FUNCTION_BLOCK "Connect"   // FB11, SCL
{ S7_Optimized_Access := 'TRUE' }
VERSION : 0.1
   VAR_INPUT
      tcon_param : TCON_Param;
   END_VAR
   VAR_IN_OUT
      requests : "Connection_Requests.UDT";
      saved_status : "Connection_Status.UDT";
   END_VAR
   VAR
      busy_delay_timer : TOF_TIME;
      error_timer : TOF_TIME;
      status_timer : TOF_TIME;
      TCON : TCON;
   END_VAR
   VAR_TEMP
      _block_status : "Connection_Status.UDT";
   END_VAR
BEGIN
   #TCON(REQ := #requests.connect,
         ID := #tcon_param.ID,
         DONE => #_block_status.done,
         BUSY => #_block_status.busy,
         ERROR => #_block_status.error,
         STATUS => #_block_status.status,
         CONNECT := #tcon_param);
   #requests.connect := FALSE;
   "Connect_Status.to_Control_Element"(requests := #requests,
                                          block_status := #_block_status,
                                          busy_timer := #busy_delay_timer,
                                          error_timer := #error_timer,
                                          saved_status := #saved_status,
                                          status_timer := #status_timer);
END_FUNCTION_BLOCK

// folder: tcpip_connection/connect/connect_status

FUNCTION "Connect_Status.Done" : Void   // FC138, SCL
{ S7_Optimized_Access := 'TRUE' }
VERSION : 0.1
   VAR_INPUT
      requests : "Connection_Requests.UDT";
      block_status : "Connection_Status.UDT";
   END_VAR
   VAR_IN_OUT
      saved_status : "Connection_Status.UDT";
   END_VAR
BEGIN
   "Connect_Status.Set_Done"(block_status := #block_status,
                                requests := #requests,
                                saved_status := #saved_status);
   "Connect_Status.Reset_Done"(block_status := #block_status,
                                  requests := #requests,
                                  saved_status := #saved_status);
END_FUNCTION

FUNCTION "Connect_Status.Error" : Void   // FC139, SCL
{ S7_Optimized_Access := 'TRUE' }
VERSION : 0.1
   VAR_INPUT
      block_status : "Connection_Status.UDT";
      requests : "Connection_Requests.UDT";
   END_VAR
   VAR_IN_OUT
      off_delay : TOF_TIME;
      saved_status : "Connection_Status.UDT";
   END_VAR
BEGIN
   "Connect_Status.Set_Error"(block_status := #block_status,
                                 requests := #requests,
                                 off_delay := #off_delay,
                                 saved_status := #saved_status);
END_FUNCTION

FUNCTION "Connect_Status.Reset_Busy" : Void   // FC140, SCL
{ S7_Optimized_Access := 'TRUE' }
VERSION : 0.1
   VAR_INPUT
      requests : "Connection_Requests.UDT";
   END_VAR
   VAR_IN_OUT
      saved_status : "Connection_Status.UDT";
   END_VAR
BEGIN
   IF #requests.disconnect THEN
       #saved_status.busy := FALSE;
   END_IF;
END_FUNCTION

FUNCTION "Connect_Status.Set_Busy" : Void   // FC142, SCL
{ S7_Optimized_Access := 'TRUE' }
VERSION : 0.1
   VAR_INPUT
      block_status : "Connection_Status.UDT";
      requests : "Connection_Requests.UDT";
   END_VAR
   VAR_IN_OUT
      off_delay : TOF_TIME;
      saved_status : "Connection_Status.UDT";
   END_VAR
   VAR_TEMP
      _et : Time;
   END_VAR
   VAR CONSTANT
      DELAY : Time := t#3s;
   END_VAR
BEGIN
   #off_delay(IN := #block_status.busy AND NOT #requests.disconnect,
              PT := #DELAY,
              Q => #saved_status.busy,
              ET => #_et);
END_FUNCTION

FUNCTION "Connect_Status.Busy" : Void   // FC143, SCL
{ S7_Optimized_Access := 'TRUE' }
VERSION : 0.1
   VAR_INPUT
      block_status : "Connection_Status.UDT";
      requests : "Connection_Requests.UDT";
   END_VAR
   VAR_IN_OUT
      off_delay : TOF_TIME;
      saved_status : "Connection_Status.UDT";
   END_VAR
BEGIN
   "Connect_Status.Set_Busy"(block_status := #block_status,
                                requests := #requests,
                                off_delay := #off_delay,
                                saved_status := #saved_status);
   "Connect_Status.Reset_Busy"(requests := #requests,
                                  saved_status := #saved_status);
END_FUNCTION

FUNCTION "Connect_Status.to_Control_Element" : Void   // FC144, SCL
{ S7_Optimized_Access := 'TRUE' }
VERSION : 0.1
   VAR_INPUT
      requests : "Connection_Requests.UDT";
      block_status : "Connection_Status.UDT";
   END_VAR
   VAR_IN_OUT
      busy_timer : TOF_TIME;
      error_timer : TOF_TIME;
      saved_status : "Connection_Status.UDT";
      status_timer : TOF_TIME;
   END_VAR
BEGIN
   "Connect_Status.Busy"(block_status := #block_status,
                            requests := #requests,
                            off_delay := #busy_timer,
                            saved_status := #saved_status);
   "Connect_Status.Done"(requests := #requests,
                            block_status := #block_status,
                            saved_status := #saved_status);
   "Connect_Status.Error"(block_status := #block_status,
                             requests := #requests,
                             off_delay := #error_timer,
                             saved_status := #saved_status);
   "Connect_Status.Status"(block_status := #block_status,
                              requests := #requests,
                              saved_status := #saved_status,
                              status_timer := #status_timer);
END_FUNCTION

FUNCTION "Connect_Status.Set_Done" : Void   // FC145, SCL
{ S7_Optimized_Access := 'TRUE' }
VERSION : 0.1
   VAR_INPUT
      block_status : "Connection_Status.UDT";
      requests : "Connection_Requests.UDT";
   END_VAR
   VAR_IN_OUT
      saved_status : "Connection_Status.UDT";
   END_VAR
BEGIN
   IF #block_status.done THEN
       #saved_status.done := TRUE;
   END_IF;
END_FUNCTION

FUNCTION "Connect_Status.Reset_Done" : Void   // FC146, SCL
{ S7_Optimized_Access := 'TRUE' }
VERSION : 0.1
   VAR_INPUT
      block_status : "Connection_Status.UDT";
      requests : "Connection_Requests.UDT";
   END_VAR
   VAR_IN_OUT
      saved_status : "Connection_Status.UDT";
   END_VAR
BEGIN
   IF #requests.disconnect THEN
       #saved_status.done := FALSE;
   END_IF;
END_FUNCTION

FUNCTION "Connect_Status.Set_Error" : Void   // FC147, SCL
{ S7_Optimized_Access := 'TRUE' }
VERSION : 0.1
   VAR_INPUT
      block_status : "Connection_Status.UDT";
      requests : "Connection_Requests.UDT";
   END_VAR
   VAR_IN_OUT
      off_delay : TOF_TIME;
      saved_status : "Connection_Status.UDT";
   END_VAR
   VAR_TEMP
      _et : Time;
   END_VAR
   VAR CONSTANT
      DELAY : Time := t#30s;
   END_VAR
BEGIN
   #off_delay(IN := #block_status.error,
              PT := #DELAY,
              Q => #saved_status.error,
              ET => #_et);
END_FUNCTION

FUNCTION "Connect_Status.Save_Status" : Void   // FC148, SCL
{ S7_Optimized_Access := 'TRUE' }
VERSION : 0.1
   VAR_INPUT
      block_status : "Connection_Status.UDT";
   END_VAR
   VAR_IN_OUT
      saved_status : "Connection_Status.UDT";
      status_timer : TOF_TIME;
   END_VAR
   VAR_TEMP
      _delay_update : Bool;
      _et : Time;
   END_VAR
   VAR CONSTANT
      DELAY : Time := T#30S;
      IDLE : Word := 16#7000;
   END_VAR
BEGIN
   IF #block_status.status <> #IDLE THEN
       #saved_status.status := #block_status.status;
   END_IF;
   #status_timer(IN := #block_status.status <> #IDLE,
                 PT := #DELAY,
                 Q => #_delay_update,
                 ET => #_et);
   IF #_delay_update THEN
       RETURN;
   END_IF;
   #saved_status.status := #block_status.status;
END_FUNCTION

FUNCTION "Connect_Status.Status" : Void   // FC149, SCL
{ S7_Optimized_Access := 'TRUE' }
VERSION : 0.1
   VAR_INPUT
      block_status : "Connection_Status.UDT";
      requests : "Connection_Requests.UDT";
   END_VAR
   VAR_IN_OUT
      saved_status : "Connection_Status.UDT";
      status_timer : TOF_TIME;
   END_VAR
BEGIN
   "Connect_Status.Save_Status"(block_status := #block_status,
                                   saved_status := #saved_status,
                                   status_timer := #status_timer);
   "Connect_Status.Clear_Status"(requests := #requests,
                                    saved_status := #saved_status);
END_FUNCTION

FUNCTION "Connect_Status.Clear_Status" : Void   // FC150, SCL
{ S7_Optimized_Access := 'TRUE' }
VERSION : 0.1
   VAR_INPUT
      requests : "Connection_Requests.UDT";
   END_VAR
   VAR_IN_OUT
      saved_status : "Connection_Status.UDT";
   END_VAR
BEGIN
   IF #requests.disconnect THEN
       #saved_status.status := 0;
   END_IF;
END_FUNCTION

// folder: tcpip_connection/connection_control

FUNCTION "Connection_Control.Initialize_Display" : Void   // FC85, SCL
{ S7_Optimized_Access := 'TRUE' }
VERSION : 0.1
   VAR_IN_OUT
      interface : "Connection_Status.HMI.UDT";
   END_VAR
BEGIN
   "Screen_Background.Initialize_Color"(#interface.background);
   "Screen_Background.Initialize_Visibility"(#interface.background);
   "Connection_Control_Table.Initialize_Display"(#interface.wire);
   "Connection_Control_Table.Initialize_Display"(#interface.material);
END_FUNCTION

// folder: tcpip_connection/connection_control/connection_control_element

FUNCTION "Connection_Control_Element.Initialize_Display" : Void   // FC86, SCL
{ S7_Optimized_Access := 'TRUE' }
VERSION : 0.1
   VAR_IN_OUT
      connection_status_element : "Connection_Status_Element.UDT";
   END_VAR
BEGIN
   "Connection_Control_Element.Initialize_Colors"(#connection_status_element);
   "Connection_Control_Element.Initialize_Visible"(#connection_status_element);
   "Connection_Control_Element.Initialize_Enable"(#connection_status_element);
END_FUNCTION

FUNCTION "Connection_Control_Element.Initialize_Colors" : Void   // FC87, SCL
{ S7_Optimized_Access := 'TRUE' }
VERSION : 0.1
   VAR_IN_OUT
      connection_status_element : "Connection_Status_Element.UDT";
   END_VAR
BEGIN
   #connection_status_element.busy_status_indicator_animate := "Color.String_to_DInt"("BUSY_INDICATOR_OFF");
   #connection_status_element.done_status_indicator_animate := "Color.String_to_DInt"("DONE_INDICATOR_OFF");
   #connection_status_element.error_status_indicator_animate := "Color.String_to_DInt"("ERROR_INDICATOR_OFF");
   #connection_status_element.operation_label_animate := "Color.String_to_DInt"("OPERATION_LABEL_OFF");
   #connection_status_element.status_code_description_animate := "Color.String_to_DInt"("STATUS_CODE_OFF");
   #connection_status_element.status_code_label_animate := "Color.String_to_DInt"("STATUS_CODE_OFF");
   #connection_status_element.status_code_value_animate := "Color.String_to_DInt"("STATUS_CODE_OFF");
END_FUNCTION

FUNCTION "Connection_Control_Element.Initialize_Visible" : Void   // FC88, SCL
{ S7_Optimized_Access := 'TRUE' }
VERSION : 0.1
   VAR_IN_OUT
      connection_status_element : "Connection_Status_Element.UDT";
   END_VAR
BEGIN
   #connection_status_element.busy_status_indicator_visible := TRUE;
   #connection_status_element.done_status_indicator_visible := TRUE;
   #connection_status_element.error_status_indicator_visible := TRUE;
   #connection_status_element.operation_button_visible := TRUE;
   #connection_status_element.operation_label_visible := TRUE;
   #connection_status_element.show_status_code_description_button_visible := TRUE;
   #connection_status_element.status_code_description_visible := TRUE;
   #connection_status_element.status_code_label_visible := TRUE;
   #connection_status_element.status_code_value_visible := TRUE;
END_FUNCTION

FUNCTION "Connection_Control_Element.Initialize_Enable" : Void   // FC89, SCL
{ S7_Optimized_Access := 'TRUE' }
VERSION : 0.1
   VAR_IN_OUT
      connection_status_element : "Connection_Status_Element.UDT";
   END_VAR
BEGIN
   #connection_status_element.operation_button_enable := TRUE;
   #connection_status_element.show_status_code_description_button_enable := TRUE;
END_FUNCTION

FUNCTION "Connection_Control_Element.Animate_Done" : Void   // FC94, SCL
{ S7_Optimized_Access := 'TRUE' }
VERSION : 0.1
   VAR_INPUT
      status : "Connection_Status.UDT";
   END_VAR
   VAR_IN_OUT
      interface : "Connection_Status_Element.UDT";
   END_VAR
BEGIN
   "Bool.Animate"(signal := #status.done,
                  color_on := "Color.String_to_DInt"("DONE_INDICATOR_ON"),
                  color_off := "Color.String_to_DInt"("DONE_INDICATOR_OFF"),
                  animation := #interface.done_status_indicator_animate);
END_FUNCTION

FUNCTION "Connection_Control_Element.Animate_Error" : Void   // FC95, SCL
{ S7_Optimized_Access := 'TRUE' }
VERSION : 0.1
   VAR_INPUT
      status : "Connection_Status.UDT";
   END_VAR
   VAR_IN_OUT
      interface : "Connection_Status_Element.UDT";
   END_VAR
BEGIN
   "Bool.Animate"(signal := #status.error,
                  color_on := "Color.String_to_DInt"("ERROR_INDICATOR_ON"),
                  color_off := "Color.String_to_DInt"("ERROR_INDICATOR_OFF"),
                  animation := #interface.error_status_indicator_animate);
END_FUNCTION

FUNCTION "Connection_Control_Element.Animate_Status_Bad" : Void   // FC96, SCL
{ S7_Optimized_Access := 'TRUE' }
VERSION : 0.1
   VAR_IN_OUT
      connection_status_element : "Connection_Status_Element.UDT";
   END_VAR
BEGIN
   #connection_status_element.status_code_description_animate := "Color.String_to_DInt"("STATUS_CODE_PROBLEM");
   #connection_status_element.status_code_label_animate := "Color.String_to_DInt"("STATUS_CODE_PROBLEM");
   #connection_status_element.status_code_value_animate := "Color.String_to_DInt"("STATUS_CODE_PROBLEM");
END_FUNCTION

FUNCTION "Connection_Control_Element.Animate_Busy" : Void   // FC97, SCL
{ S7_Optimized_Access := 'TRUE' }
VERSION : 0.1
   VAR_INPUT
      status : "Connection_Status.UDT";
   END_VAR
   VAR_IN_OUT
      element : "Connection_Status_Element.UDT";
   END_VAR
BEGIN
   "Bool.Animate"(signal := #status.busy,
                  color_on := "Color.String_to_DInt"("BUSY_INDICATOR_ON"),
                  color_off := "Color.String_to_DInt"("BUSY_INDICATOR_OFF"),
                  animation := #element.busy_status_indicator_animate);
END_FUNCTION

FUNCTION "Connection_Control_Element.Animate_Status_Good" : Void   // FC98, SCL
{ S7_Optimized_Access := 'TRUE' }
VERSION : 0.1
   VAR_IN_OUT
      interface : "Connection_Status_Element.UDT";
   END_VAR
BEGIN
   #interface.status_code_description_animate := "Color.String_to_DInt"("STATUS_CODE_GOOD");
   #interface.status_code_label_animate := "Color.String_to_DInt"("STATUS_CODE_GOOD");
   #interface.status_code_value_animate := "Color.String_to_DInt"("STATUS_CODE_GOOD");
END_FUNCTION

FUNCTION "Connection_Control_Element.Animate_Operation_Acutate" : Void   // FC135, SCL
{ S7_Optimized_Access := 'TRUE' }
VERSION : 0.1
   VAR_IN_OUT
      interface : "Connection_Status_Element.UDT";
   END_VAR
   VAR_TEMP
      _animation : DInt;
   END_VAR
BEGIN
   "Bool.Animate"(signal := #interface.operation_button_actuate,
                  color_on := "Color.String_to_DInt"("ACTUATE"),
                  color_off := "Color.String_to_DInt"("OPERATION_OFF"),
                  animation := #interface.operation_label_animate);
END_FUNCTION

FUNCTION "Connection_Control_Element.Animate" : Void   // FC141, SCL
{ S7_Optimized_Access := 'TRUE' }
VERSION : 0.1
   VAR_INPUT
      status : "Connection_Status.UDT";
   END_VAR
   VAR_IN_OUT
      interface : "Connection_Status_Element.UDT";
   END_VAR
BEGIN
   "Connection_Control_Element.Animate_Operation_Acutate"(#interface);
   "Connection_Control_Element.Animate_Busy"(status := #status,
                                             element := #interface);
   "Connection_Control_Element.Animate_Done"(status := #status,
                                             interface := #interface);
   "Connection_Control_Element.Animate_Error"(status := #status,
                                              interface := #interface);
   "Connection_Status_Element.Animate_Status"(status := #status,
                                              interface := #interface);
END_FUNCTION

FUNCTION "Connection_Status_Element.Animate_Status" : Void   // FC151, SCL
{ S7_Optimized_Access := 'TRUE' }
VERSION : 0.1
   VAR_INPUT
      status : "Connection_Status.UDT";
   END_VAR
   VAR_IN_OUT
      interface : "Connection_Status_Element.UDT";
   END_VAR
BEGIN
   #interface.status_code_description_value := WORD_TO_DINT(#status.status);
   #interface.status_code_value := "Word.to_String"(#status.status);
   CASE #status.status OF
       "IDLE", "SUCCESS":
           "Connection_Control_Element.Animate_Status_Good"(#interface);
       ELSE
           "Connection_Control_Element.Animate_Status_Bad"(#interface);
   END_CASE;
END_FUNCTION

// folder: tcpip_connection/connection_control/connection_control_header

FUNCTION "Connection_Control_Header.Initialize_Display" : Void   // FC91, SCL
{ S7_Optimized_Access := 'TRUE' }
VERSION : 0.1
   VAR_IN_OUT
      interface : "Connection_Status_Header.UDT";
   END_VAR
BEGIN
   "Connection_Control_Header.Initialize_Color"(#interface);
   "Connection_Control_Header.Initialize_Visible"(#interface);
   "Connection_Control_Header.Initialize_Enable"(#interface);
END_FUNCTION

FUNCTION "Connection_Control_Header.Initialize_Color" : Void   // FC92, SCL
{ S7_Optimized_Access := 'TRUE' }
VERSION : 0.1
   VAR_IN_OUT
      connection_status_header : "Connection_Status_Header.UDT";
   END_VAR
BEGIN
   #connection_status_header.animate := "Color.String_to_DInt"("CONNECTION_STATUS_HEADER");
END_FUNCTION

FUNCTION "Connection_Control_Header.Initialize_Visible" : Void   // FC93, SCL
{ S7_Optimized_Access := 'TRUE' }
VERSION : 0.1
   VAR_IN_OUT
      connection_status_header : "Connection_Status_Header.UDT";
   END_VAR
BEGIN
   #connection_status_header.visible := TRUE;
END_FUNCTION

FUNCTION "Connection_Control_Header.Initialize_Enable" : Void   // FC107, SCL
{ S7_Optimized_Access := 'TRUE' }
VERSION : 0.1
   VAR_IN_OUT
      interface : "Connection_Status_Header.UDT";
   END_VAR
BEGIN
   #interface.enable := TRUE;
END_FUNCTION

FUNCTION "Connection_Control.Animate_Header" : Void   // FC129, SCL
{ S7_Optimized_Access := 'TRUE' }
VERSION : 0.1
   VAR_IN_OUT
      interface : "Connection_Status_Header.UDT";
   END_VAR
BEGIN
   "Bool.Animate"(signal := #interface.actuate,
                  color_on := "Color.String_to_DInt"("ACTUATE"),
                  color_off := "Color.String_to_DInt"("LABEL_COLOR"),
                  animation := #interface.animate);
END_FUNCTION

// folder: tcpip_connection/connection_control/connection_control_table

FUNCTION "Connection_Control_Table.Initialize_Display" : Void   // FC90, SCL
{ S7_Optimized_Access := 'TRUE' }
VERSION : 0.1
   VAR_IN_OUT
      connection_status_table : "Connection_Status_Table.UDT";
   END_VAR
BEGIN
   "Connection_Control_Header.Initialize_Display"(#connection_status_table.header);
   "Connection_Control_Element.Initialize_Display"(#connection_status_table.disconnect);
   "Connection_Control_Element.Initialize_Display"(#connection_status_table.connect);
   "Connection_Control_Element.Initialize_Display"(#connection_status_table.send);
END_FUNCTION

FUNCTION "Connection_Control_Table.Animate" : Void   // FC136, SCL
{ S7_Optimized_Access := 'TRUE' }
VERSION : 0.1
   VAR_INPUT
      statuses : "Connection_Statuses.UDT";
   END_VAR
   VAR_IN_OUT
      interface : "Connection_Status_Table.UDT";
   END_VAR
BEGIN
   "Connection_Control.Animate_Header"(#interface.header);
   "Connection_Control_Element.Animate"(status := #statuses.connect,
                                        interface := #interface.connect);
   "Connection_Control_Element.Animate"(status := #statuses.disconnect,
                                        interface := #interface.disconnect);
   "Connection_Control_Element.Animate"(status := #statuses.send,
                                        interface := #interface.send);
END_FUNCTION

// folder: tcpip_connection/connection_parameters

FUNCTION "Connection_Parameters.Initialize_Colors" : Void   // FC108, SCL
{ S7_Optimized_Access := 'TRUE' }
VERSION : 0.1
   VAR_IN_OUT
      interface : "Connection_Parameters_HMI_Interface.UDT";
   END_VAR
BEGIN
   #interface.back_animate := "Color.String_to_DInt"("LABEL_COLOR");
   #interface.header_animate := "Color.String_to_DInt"("LABEL_COLOR");
   #interface.id_entry_animate := "Color.String_to_DInt"("DESELECTED_INPUT_COLOR");
   #interface.id_label_animate := "Color.String_to_DInt"("LABEL_COLOR");
   #interface.ip_address_entry_animate := "Color.String_to_DInt"("DESELECTED_INPUT_COLOR");
   #interface.ip_address_label_animate := "Color.String_to_DInt"("LABEL_COLOR");
   #interface.port_entry_animate := "Color.String_to_DInt"("DESELECTED_INPUT_COLOR");
   #interface.port_label_animate := "Color.String_to_DInt"("LABEL_COLOR");
   #interface.back_animate := "Color.String_to_DInt"("LABEL_COLOR");
END_FUNCTION

FUNCTION "Connection_Parameters.Initialize_Visible" : Void   // FC109, SCL
{ S7_Optimized_Access := 'TRUE' }
VERSION : 0.1
   VAR_IN_OUT
      interface : "Connection_Parameters_HMI_Interface.UDT";
   END_VAR
BEGIN
   #interface.back_visible := TRUE;
   #interface.header_visible := TRUE;
   #interface.id_entry_visible := TRUE;
   #interface.id_label_visible := TRUE;
   #interface.ip_address_entry_visible := TRUE;
   #interface.ip_address_label_visible := TRUE;
   #interface.port_entry_visible := TRUE;
   #interface.port_label_visible := TRUE;
END_FUNCTION

FUNCTION "Connection_Parameters.Initialize_Enable" : Void   // FC110, SCL
{ S7_Optimized_Access := 'TRUE' }
VERSION : 0.1
   VAR_IN_OUT
      interface : "Connection_Parameters_HMI_Interface.UDT";
   END_VAR
BEGIN
   #interface.back_enable := TRUE;
   #interface.id_entry_enable := TRUE;
   #interface.ip_address_entry_enable := TRUE;
   #interface.port_entry_enable := TRUE;
   #interface.back_enable := TRUE;
END_FUNCTION

FUNCTION "Connection_Parameters.Initialize_Display" : Void   // FC111, SCL
{ S7_Optimized_Access := 'TRUE' }
VERSION : 0.1
   VAR_IN_OUT
      interface : "Connection_Paramters_HMI.UDT";
   END_VAR
BEGIN
   "Screen_Background.Initialize"(#interface.background);
   "Connection_Parameters.Initialize_Controls_Display"(#interface.connection_parameters);
END_FUNCTION

FUNCTION "Connection_Parameters.Initialize_Controls_Display" : Void   // FC112, SCL
{ S7_Optimized_Access := 'TRUE' }
VERSION : 0.1
   VAR_IN_OUT
      interface : "Connection_Parameters_HMI_Interface.UDT";
   END_VAR
BEGIN
   "Connection_Parameters.Initialize_Colors"(#interface);
   "Connection_Parameters.Initialize_Visible"(#interface);
   "Connection_Parameters.Initialize_Enable"(#interface);
END_FUNCTION

FUNCTION "Connection_Parameters.Make_Header_Text" : Void   // FC113, SCL
{ S7_Optimized_Access := 'TRUE' }
VERSION : 0.1
   VAR_INPUT
      "name" : String;
   END_VAR
   VAR_IN_OUT
      interface : "Connection_Parameters_HMI_Interface.UDT";
   END_VAR
BEGIN
   #interface.header_value := CONCAT_STRING(IN1 := #name,
                                            IN2 := ' PARAMETERS');
END_FUNCTION

FUNCTION "Connection_Parameters.Get_Parameters" : Void   // FC114, SCL
{ S7_Optimized_Access := 'TRUE' }
VERSION : 0.1
   VAR_INPUT
      connection_parameters : "Connection_Parameters.UDT";
   END_VAR
   VAR_IN_OUT
      interface : "Connection_Parameters_HMI_Interface.UDT";
   END_VAR
BEGIN
   #interface.id_entry_value := "Word.to_String"(#connection_parameters.id);
   #interface.ip_address_entry_value := #connection_parameters.ip_address;
   #interface.port_entry_value := #connection_parameters.port_number;
END_FUNCTION

FUNCTION "Connection_Parameters.Set_ID" : Void   // FC115, SCL
{ S7_Optimized_Access := 'TRUE' }
VERSION : 0.1
   VAR_INPUT
      interface : "Connection_Parameters_HMI_Interface.UDT";
   END_VAR
   VAR_IN_OUT
      connection_parameters : "Connection_Parameters.UDT";
   END_VAR
BEGIN
   IF NOT "Connection_Parameters.ID_Is_Valid"(#interface.id_entry_value) THEN
       RETURN;
   END_IF;
   #connection_parameters.id := UINT_TO_WORD(STRING_TO_UINT(#interface.id_entry_value));
   RETURN;
END_FUNCTION

FUNCTION "Connection_Parameters.IP_Address_Is_Valid" : Bool   // FC119, SCL
{ S7_Optimized_Access := 'TRUE' }
VERSION : 0.1
   VAR_INPUT
      ip_address : String;
   END_VAR
BEGIN
   IF FIND(IN1 := #ip_address, IN2 := '.') > 0 THEN
       #"Connection_Parameters.IP_Address_Is_Valid" := TRUE;
       RETURN;
   END_IF;
   IF FIND(IN1 := #ip_address, IN2 := '_') > 0 THEN
       #"Connection_Parameters.IP_Address_Is_Valid" := TRUE;
       RETURN;
   END_IF;
   #"Connection_Parameters.IP_Address_Is_Valid" := FALSE;
   RETURN;
END_FUNCTION

FUNCTION "Connection_Parameters.Set_Parameters" : Void   // FC120, SCL
{ S7_Optimized_Access := 'TRUE' }
VERSION : 0.1
   VAR_IN_OUT
      interface : "Connection_Parameters_HMI_Interface.UDT";
      saved : "Connection_Parameters.UDT";
   END_VAR
BEGIN
   IF #interface.id_entry_input_finished THEN
       #interface.id_entry_input_finished := FALSE;
       "Connection_Parameters.Set_ID"(interface := #interface,
                                      connection_parameters := #saved);
       RETURN;
   END_IF;
   IF #interface.ip_address_entry_input_finished THEN
       #interface.ip_address_entry_input_finished := FALSE;
       "Connection_Parameters.Set_IP_Address"(interface := #interface,
                                              connection_parameters := #saved);
       RETURN;
   END_IF;
   IF #interface.port_entry_input_finished THEN
       #interface.port_entry_input_finished := FALSE;
       "Connection_Parameters.Set_Port"(interface := #interface,
                                        connection_parameters := #saved);
       RETURN;
   END_IF;
END_FUNCTION

FUNCTION "Connection_Parameters.Set_Mode" : Void   // FC121, SCL
{ S7_Optimized_Access := 'TRUE' }
VERSION : 0.1
   VAR_INPUT
      interface : "Connection_Status.HMI.UDT";
   END_VAR
   VAR_IN_OUT
      meta : "HMI_Meta.UDT";
   END_VAR
BEGIN
   IF #interface.material.header.actuate THEN
       #meta.parameter_entry_mode := "MATERIAL";
   END_IF;
   IF #interface.wire.header.actuate THEN
       #meta.parameter_entry_mode := "WIRE";
   END_IF;
END_FUNCTION

FUNCTION "Connection_Parameters.Reload_Screen" : Void   // FC122, SCL
{ S7_Optimized_Access := 'TRUE' }
VERSION : 0.1
   VAR_INPUT
      meta : "HMI_Meta.UDT";
      connection_controls : "Connection_Status.HMI.UDT";
      led : "LED_Interfaces.UDT";
   END_VAR
   VAR_IN_OUT
      hmi : "Connection_Paramters_HMI.UDT";
   END_VAR
BEGIN
   "Connection_Parameters.Make_Header_Text"(name := #meta.parameter_entry_mode,
                                            interface := #hmi.connection_parameters);
   IF #meta.parameter_entry_mode = "MATERIAL" THEN
       "Connection_Parameters.Get_Parameters"(connection_parameters := #led.material.connection_parameters,
                                              interface := #hmi.connection_parameters);
   END_IF;
   IF #meta.parameter_entry_mode = "WIRE" THEN
       "Connection_Parameters.Get_Parameters"(connection_parameters := #led.wire.connection_parameters,
                                              interface := #hmi.connection_parameters);
   END_IF;
END_FUNCTION

FUNCTION "Connection_Parameters.Set_IP_Address" : Void   // FC124, SCL
{ S7_Optimized_Access := 'TRUE' }
VERSION : 0.1
   VAR_INPUT
      interface : "Connection_Parameters_HMI_Interface.UDT";
   END_VAR
   VAR_IN_OUT
      connection_parameters : "Connection_Parameters.UDT";
   END_VAR
BEGIN
   IF NOT "Connection_Parameters.IP_Address_Is_Valid"(#interface.ip_address_entry_value) THEN
       RETURN;
   END_IF;
   #connection_parameters.ip_address := #interface.ip_address_entry_value;
   RETURN;
END_FUNCTION

FUNCTION "Connection_Parameters.Set_Port" : Void   // FC125, SCL
{ S7_Optimized_Access := 'TRUE' }
VERSION : 0.1
   VAR_INPUT
      interface : "Connection_Parameters_HMI_Interface.UDT";
   END_VAR
   VAR_IN_OUT
      connection_parameters : "Connection_Parameters.UDT";
   END_VAR
BEGIN
   IF NOT "Connection_Parameters.Port_Is_Valid"(#interface.port_entry_value) THEN
       RETURN;
   END_IF;
   #connection_parameters.port_number := #interface.port_entry_value;
   RETURN;
END_FUNCTION

FUNCTION "Connection_Parameters.Port_Is_Valid" : Bool   // FC126, SCL
{ S7_Optimized_Access := 'TRUE' }
VERSION : 0.1
   VAR_INPUT
      port : String;
   END_VAR
BEGIN
   IF "String.Is_Numeric"(#port) THEN
       #"Connection_Parameters.Port_Is_Valid" := TRUE;
       RETURN;
   END_IF;
   #"Connection_Parameters.Port_Is_Valid" := FALSE;
   RETURN;
END_FUNCTION

FUNCTION "Connection_Parameters.ID_Is_Valid" : Bool   // FC127, SCL
{ S7_Optimized_Access := 'TRUE' }
VERSION : 0.1
   VAR_INPUT
      id : String;
   END_VAR
BEGIN
   IF "String.Is_Numeric"(#id) THEN
       #"Connection_Parameters.ID_Is_Valid" := TRUE;
       RETURN;
   END_IF;
   #"Connection_Parameters.ID_Is_Valid" := FALSE;
   RETURN;
END_FUNCTION

FUNCTION "Connection_Parameters.Animate_Back" : Void   // FC130, SCL
{ S7_Optimized_Access := 'TRUE' }
VERSION : 0.1
   VAR_IN_OUT
      interface : "Connection_Parameters_HMI_Interface.UDT";
   END_VAR
BEGIN
   "Bool.Animate"(signal := #interface.back_actuate,
                  color_on := "Color.String_to_DInt"("ACTUATE"),
                  color_off := "Color.String_to_DInt"("LABEL_COLOR"),
                  animation := #interface.back_animate);
END_FUNCTION

FUNCTION "Connection_Parameters.Animate_ID_Active" : Void   // FC132, SCL
{ S7_Optimized_Access := 'TRUE' }
VERSION : 0.1
   VAR_IN_OUT
      interface : "Connection_Parameters_HMI_Interface.UDT";
   END_VAR
BEGIN
   "Bool.Animate"(signal := #interface.id_entry_active,
                  color_on := "Color.String_to_DInt"("SELECTED_INPUT_COLOR"),
                  color_off := "Color.String_to_DInt"("DESELECTED_INPUT_COLOR"),
                  animation := #interface.id_entry_animate);
END_FUNCTION

FUNCTION "Connection_Parameters.Animate_Port_Active" : Void   // FC133, SCL
{ S7_Optimized_Access := 'TRUE' }
VERSION : 0.1
   VAR_IN_OUT
      interface : "Connection_Parameters_HMI_Interface.UDT";
   END_VAR
BEGIN
   "Bool.Animate"(signal := #interface.port_entry_active,
                  color_on := "Color.String_to_DInt"("SELECTED_INPUT_COLOR"),
                  color_off := "Color.String_to_DInt"("DESELECTED_INPUT_COLOR"),
                  animation := #interface.port_entry_animate);
END_FUNCTION

FUNCTION "Connection_Parameters.Animate_IP_Active" : Void   // FC134, SCL
{ S7_Optimized_Access := 'TRUE' }
VERSION : 0.1
   VAR_IN_OUT
      interface : "Connection_Parameters_HMI_Interface.UDT";
   END_VAR
BEGIN
   "Bool.Animate"(signal := #interface.ip_address_entry_active,
                  color_on := "Color.String_to_DInt"("SELECTED_INPUT_COLOR"),
                  color_off := "Color.String_to_DInt"("DESELECTED_INPUT_COLOR"),
                  animation := #interface.ip_address_entry_animate);
END_FUNCTION

// folder: tcpip_connection/connection_status_details

FUNCTION "Connection_Status_Details.Initialize_Display" : Void   // FC165, SCL
{ S7_Optimized_Access := 'TRUE' }
VERSION : 0.1
   VAR_IN_OUT
      interface : "Connection_Detail.HMI.UDT";
   END_VAR
BEGIN
   "Connection_Status_Details.Initialize_Colors"(#interface);
   "Connection_Status_Details.Initialize_Enable"(#interface);
   "Connection_Status_Details.Initialize_Visible"(#interface);
END_FUNCTION

FUNCTION "Connection_Status_Details.Initialize_Visible" : Void   // FC184, SCL
{ S7_Optimized_Access := 'TRUE' }
VERSION : 0.1
   VAR_IN_OUT
      interface : "Connection_Detail.HMI.UDT";
   END_VAR
BEGIN
   #interface.back_button_visible := TRUE;
   #interface.detailed_status_visible := TRUE;
   #interface.display_payload_button_visible := TRUE;
   #interface.header_visible := true;
   #interface.payload_visible := TRUE;
END_FUNCTION

FUNCTION "Connection_Status_Details.Initialize_Colors" : Void   // FC185, SCL
{ S7_Optimized_Access := 'TRUE' }
VERSION : 0.1
   VAR_IN_OUT
      interface : "Connection_Detail.HMI.UDT";
   END_VAR
BEGIN
   #interface.detailed_status_animate := "Color.String_to_DInt"("LABEL_COLOR");
   #interface.display_payload_button_animate := "Color.String_to_DInt"("LABEL_COLOR");
   #interface.header_animate := "Color.String_to_DInt"("LABEL_COLOR");
   #interface.payload_animate := "Color.String_to_DInt"("LABEL_COLOR");
END_FUNCTION

FUNCTION "Connection_Status_Details.Initialize_Enable" : Void   // FC186, SCL
{ S7_Optimized_Access := 'TRUE' }
VERSION : 0.1
   VAR_IN_OUT
      interface : "Connection_Detail.HMI.UDT";
   END_VAR
BEGIN
   #interface.back_button_enable := TRUE;
   #interface.display_payload_button_enable := TRUE;
END_FUNCTION

FUNCTION "Connection_Status_Details.Set_Mode" : Void   // FC187, SCL
{ S7_Optimized_Access := 'TRUE' }
VERSION : 0.1
   VAR_INPUT
      interface : "Connection_Status.HMI.UDT";
   END_VAR
   VAR_IN_OUT
      mode : DInt;
   END_VAR
BEGIN
   IF #interface.material.disconnect.show_status_code_description_button_actuate THEN
       #mode := "MATERIAL_DISCONNECT";
       RETURN;
   END_IF;

   IF #interface.material.connect.show_status_code_description_button_actuate THEN
       #mode := "MATERIAL_CONNECT";
       RETURN;
   END_IF;

   IF #interface.material.send.show_status_code_description_button_actuate THEN
       #mode := "MATERIAL_SEND";
       RETURN;
   END_IF;

   IF #interface.wire.disconnect.show_status_code_description_button_actuate THEN
       #mode := "WIRE_DISCONNECT";
       RETURN;
   END_IF;

   IF #interface.wire.connect.show_status_code_description_button_actuate THEN
       #mode := "WIRE_CONNECT";
       RETURN;
   END_IF;

   IF #interface.wire.send.show_status_code_description_button_actuate THEN
       #mode := "WIRE_SEND";
       RETURN;
   END_IF;
END_FUNCTION

FUNCTION "Connection_Status_Details.Set_Header_Selector" : Void   // FC188, SCL
{ S7_Optimized_Access := 'TRUE' }
VERSION : 0.1
   VAR_INPUT
      meta : "HMI_Meta.UDT";
   END_VAR
   VAR_IN_OUT
      interface : "Connection_Detail.HMI.UDT";
   END_VAR
BEGIN
   CASE #meta.connection_mode OF

       "MATERIAL_DISCONNECT", "WIRE_DISCONNECT":
           #interface.header_selector := "DISCONNECT_SELECTOR";

       "MATERIAL_CONNECT", "WIRE_CONNECT":
           #interface.header_selector := "CONNECT_SELECTOR";

       "MATERIAL_SEND", "WIRE_SEND":
           #interface.header_selector := "SEND_SELECTOR";

   END_CASE;
END_FUNCTION

FUNCTION "Connection_Status_Details.Animate_Header" : Void   // FC189, SCL
{ S7_Optimized_Access := 'TRUE' }
VERSION : 0.1
   VAR_INPUT
      meta : "HMI_Meta.UDT";
   END_VAR
   VAR_IN_OUT
      interface : "Connection_Detail.HMI.UDT";
   END_VAR
BEGIN
   "Connection_Status_Details.Set_Header_Selector"(meta := #meta,
                                                   interface := #interface);
END_FUNCTION

FUNCTION "Connection_Status_Details.Set_Status_Details_Selector" : Void   // FC190, SCL
{ S7_Optimized_Access := 'TRUE' }
VERSION : 0.1
   VAR_INPUT
      led_interfaces : "LED_Interfaces.UDT";
      hmi_meta : "HMI_Meta.UDT";
   END_VAR
   VAR_IN_OUT
      interface : "Connection_Detail.HMI.UDT";
   END_VAR
BEGIN
   CASE #hmi_meta.connection_mode OF

       "MATERIAL_DISCONNECT":
           #interface.detailed_status_list_selector := "DISCONNECT_SELECTOR";
           #interface.detailed_status_message_selector := WORD_TO_DINT(#led_interfaces.material.statuses.disconnect.status);

       "MATERIAL_CONNECT":
           #interface.detailed_status_list_selector := "CONNECT_SELECTOR";
           #interface.detailed_status_message_selector := WORD_TO_DINT(#led_interfaces.material.statuses.connect.status);

       "MATERIAL_SEND":
           #interface.detailed_status_list_selector := "SEND_SELECTOR";
           #interface.detailed_status_message_selector := WORD_TO_DINT(#led_interfaces.material.statuses.send.status);

       "WIRE_DISCONNECT":
           #interface.detailed_status_list_selector := "DISCONNECT_SELECTOR";
           #interface.detailed_status_message_selector := WORD_TO_DINT(#led_interfaces.wire.statuses.disconnect.status);

       "WIRE_CONNECT":
           #interface.detailed_status_list_selector := "CONNECT_SELECTOR";
           #interface.detailed_status_message_selector := WORD_TO_DINT(#led_interfaces.wire.statuses.connect.status);

       "WIRE_SEND":
           #interface.detailed_status_list_selector := "SEND_SELECTOR";
           #interface.detailed_status_message_selector := WORD_TO_DINT(#led_interfaces.wire.statuses.send.status);

   END_CASE;
END_FUNCTION

FUNCTION "Connection_Status_Details.Show_Payload" : Void   // FC191, SCL
{ S7_Optimized_Access := 'TRUE' }
VERSION : 0.1
   VAR_INPUT
      led_interfaces : "LED_Interfaces.UDT";
      hmi_meta : "HMI_Meta.UDT";
   END_VAR
   VAR_IN_OUT
      interface : "Connection_Detail.HMI.UDT";
   END_VAR
   VAR_TEMP
      _delimeters : Array[0..1] of String;
      _payload_text : String;
      _send_buffer : "ADP.Message_Buffer.UDT";
   END_VAR
BEGIN
   CASE #hmi_meta.connection_mode OF

       "MATERIAL_CONNECT", "MATERIAL_DISCONNECT", "MATERIAL_SEND":  
           #_send_buffer := #led_interfaces.material.send_buffer;

       "WIRE_DISCONNECT", "WIRE_CONNECT", "WIRE_SEND":
           #_send_buffer := #led_interfaces.wire.send_buffer;

   END_CASE;

   #_payload_text := "ADP.Buffer_to_String"(buffer := #_send_buffer,
                                            lenWrap := 25);

   #_delimeters[0] := ' ';
   #_delimeters[1] := '-';
   #interface.payload_text := #_payload_text;

   #interface.payload_visible := TRUE;
   #interface.detailed_status_visible := FALSE;
END_FUNCTION

FUNCTION "Connection_Status_Details.Display_Detailed_Status" : Void   // FC193, SCL
{ S7_Optimized_Access := 'TRUE' }
VERSION : 0.1
   VAR_IN_OUT
      interface : "Connection_Detail.HMI.UDT";
   END_VAR
BEGIN
   #interface.payload_visible := FALSE;
   #interface.detailed_status_visible := TRUE;
END_FUNCTION

// folder: tcpip_connection/diagnostics

FUNCTION_BLOCK "Diagnostics"   // FB14, SCL
{ S7_Optimized_Access := 'TRUE' }
VERSION : 0.1
   VAR_INPUT
      tcon_param : TCON_Param;
   END_VAR
   VAR_IN_OUT
      requests : "Connection_Requests.UDT";
   END_VAR
   VAR
      T_DIAG : T_DIAG;
   END_VAR
BEGIN
   #T_DIAG(REQ := #requests.diagnostics,
           ID := #tcon_param.ID);
   #requests.diagnostics := FALSE;
END_FUNCTION_BLOCK

// folder: tcpip_connection/disconnect

FUNCTION_BLOCK "Disconnect"   // FB13, SCL
{ S7_Optimized_Access := 'TRUE' }
VERSION : 0.1
   VAR_INPUT
      tcon_param : TCON_Param;
   END_VAR
   VAR_IN_OUT
      requests : "Connection_Requests.UDT";
      saved_status : "Connection_Status.UDT";
   END_VAR
   VAR
      TDISCON : TDISCON;
      timers : "Connection_Status_Timers.UDT";
   END_VAR
   VAR_TEMP
      block_status : "Connection_Status.UDT";
   END_VAR
BEGIN
   #TDISCON(REQ := #requests.disconnect,
            ID := #tcon_param.ID,
            DONE => #block_status.done,
            BUSY => #block_status.busy,
            ERROR => #block_status.error,
            STATUS => #block_status.status);
   #requests.disconnect := FALSE;
   "Disconnect_Status.to_Control_Element"(requests := #requests,
                                          block_status := #block_status,
                                          saved_status := #saved_status,
                                          timers := #timers);
END_FUNCTION_BLOCK

// folder: tcpip_connection/disconnect/disconnect_status

FUNCTION "Disconnect_Status.Done" : Void   // FC152, SCL
{ S7_Optimized_Access := 'TRUE' }
VERSION : 0.1
   VAR_INPUT
      requests : "Connection_Requests.UDT";
      block_status : "Connection_Status.UDT";
   END_VAR
   VAR_IN_OUT
      saved_status : "Connection_Status.UDT";
   END_VAR
BEGIN
   "Disconnect_Status.Set_Done"(block_status := #block_status,
                                requests := #requests,
                                saved_status := #saved_status);
   "Disconnect_Status.Reset_Done"(block_status := #block_status,
                                  requests := #requests,
                                  saved_status := #saved_status);
END_FUNCTION

FUNCTION "Disconnect_Status.Error" : Void   // FC153, SCL
{ S7_Optimized_Access := 'TRUE' }
VERSION : 0.1
   VAR_INPUT
      block_status : "Connection_Status.UDT";
      requests : "Connection_Requests.UDT";
   END_VAR
   VAR_IN_OUT
      off_delay : TOF_TIME;
      saved_status : "Connection_Status.UDT";
   END_VAR
BEGIN
   "Disconnect_Status.Set_Error"(block_status := #block_status,
                                 requests := #requests,
                                 off_delay := #off_delay,
                                 saved_status := #saved_status);
END_FUNCTION

FUNCTION "Disconnect_Status.Reset_Busy" : Void   // FC154, SCL
{ S7_Optimized_Access := 'TRUE' }
VERSION : 0.1
   VAR_INPUT
      requests : "Connection_Requests.UDT";
   END_VAR
   VAR_IN_OUT
      saved_status : "Connection_Status.UDT";
   END_VAR
BEGIN
   IF #requests.connect THEN
       #saved_status.busy := FALSE;
   END_IF;
END_FUNCTION

FUNCTION "Disconnect_Status.Set_Busy" : Void   // FC155, SCL
{ S7_Optimized_Access := 'TRUE' }
VERSION : 0.1
   VAR_INPUT
      block_status : "Connection_Status.UDT";
      requests : "Connection_Requests.UDT";
   END_VAR
   VAR_IN_OUT
      off_delay : TOF_TIME;
      saved_status : "Connection_Status.UDT";
   END_VAR
   VAR_TEMP
      _et : Time;
   END_VAR
   VAR CONSTANT
      DELAY : Time := t#3s;
   END_VAR
BEGIN
   #off_delay(IN := #block_status.busy AND NOT #requests.disconnect,
              PT := #DELAY,
              Q => #saved_status.busy,
              ET => #_et);
END_FUNCTION

FUNCTION "Disconnect_Status.Busy" : Void   // FC156, SCL
{ S7_Optimized_Access := 'TRUE' }
VERSION : 0.1
   VAR_INPUT
      block_status : "Connection_Status.UDT";
      requests : "Connection_Requests.UDT";
   END_VAR
   VAR_IN_OUT
      off_delay : TOF_TIME;
      saved_status : "Connection_Status.UDT";
   END_VAR
BEGIN
   "Disconnect_Status.Set_Busy"(block_status := #block_status,
                                requests := #requests,
                                off_delay := #off_delay,
                                saved_status := #saved_status);
   "Disconnect_Status.Reset_Busy"(requests := #requests,
                                  saved_status := #saved_status);
END_FUNCTION

FUNCTION "Disconnect_Status.to_Control_Element" : Void   // FC157, SCL
{ S7_Optimized_Access := 'TRUE' }
VERSION : 0.1
   VAR_INPUT
      requests : "Connection_Requests.UDT";
      block_status : "Connection_Status.UDT";
   END_VAR
   VAR_IN_OUT
      saved_status : "Connection_Status.UDT";
      timers : "Connection_Status_Timers.UDT";
   END_VAR
BEGIN
   "Disconnect_Status.Busy"(block_status := #block_status,
                            requests := #requests,
                            off_delay := #timers.busy,
                            saved_status := #saved_status);
   "Disconnect_Status.Done"(requests := #requests,
                            block_status := #block_status,
                            saved_status := #saved_status);
   "Disconnect_Status.Error"(block_status := #block_status,
                             requests := #requests,
                             off_delay := #timers.error,
                             saved_status := #saved_status);
   "Disconnect_Status.Status"(block_status := #block_status,
                              requests := #requests,
                              saved_status := #saved_status,
                              status_timer := #timers.status);
END_FUNCTION

FUNCTION "Disconnect_Status.Set_Done" : Void   // FC158, SCL
{ S7_Optimized_Access := 'TRUE' }
VERSION : 0.1
   VAR_INPUT
      block_status : "Connection_Status.UDT";
      requests : "Connection_Requests.UDT";
   END_VAR
   VAR_IN_OUT
      saved_status : "Connection_Status.UDT";
   END_VAR
BEGIN
   IF #block_status.done THEN
       #saved_status.done := TRUE;
   END_IF;
END_FUNCTION

FUNCTION "Disconnect_Status.Reset_Done" : Void   // FC159, SCL
{ S7_Optimized_Access := 'TRUE' }
VERSION : 0.1
   VAR_INPUT
      block_status : "Connection_Status.UDT";
      requests : "Connection_Requests.UDT";
   END_VAR
   VAR_IN_OUT
      saved_status : "Connection_Status.UDT";
   END_VAR
BEGIN
   IF #requests.connect THEN
       #saved_status.done := FALSE;
   END_IF;
END_FUNCTION

FUNCTION "Disconnect_Status.Set_Error" : Void   // FC160, SCL
{ S7_Optimized_Access := 'TRUE' }
VERSION : 0.1
   VAR_INPUT
      block_status : "Connection_Status.UDT";
      requests : "Connection_Requests.UDT";
   END_VAR
   VAR_IN_OUT
      off_delay : TOF_TIME;
      saved_status : "Connection_Status.UDT";
   END_VAR
   VAR_TEMP
      _et : Time;
   END_VAR
   VAR CONSTANT
      DELAY : Time := t#30s;
   END_VAR
BEGIN
   #off_delay(IN := #block_status.error,
              PT := #DELAY,
              Q => #saved_status.error,
              ET => #_et);
END_FUNCTION

FUNCTION "Disconnect_Status.Save_Status" : Void   // FC161, SCL
{ S7_Optimized_Access := 'TRUE' }
VERSION : 0.1
   VAR_INPUT
      block_status : "Connection_Status.UDT";
   END_VAR
   VAR_IN_OUT
      saved_status : "Connection_Status.UDT";
      status_timer : TOF_TIME;
   END_VAR
   VAR_TEMP
      _delay_update : Bool;
      _et : Time;
   END_VAR
   VAR CONSTANT
      DELAY : Time := T#30S;
      IDLE : Word := 16#7000;
   END_VAR
BEGIN
   IF #block_status.status <> #IDLE THEN
       #saved_status.status := #block_status.status;
   END_IF;
   #status_timer(IN := #block_status.status <> #IDLE,
                 PT := #DELAY,
                 Q => #_delay_update,
                 ET => #_et);
   IF #_delay_update THEN
       RETURN;
   END_IF;
   #saved_status.status := #block_status.status;
END_FUNCTION

FUNCTION "Disconnect_Status.Status" : Void   // FC162, SCL
{ S7_Optimized_Access := 'TRUE' }
VERSION : 0.1
   VAR_INPUT
      block_status : "Connection_Status.UDT";
      requests : "Connection_Requests.UDT";
   END_VAR
   VAR_IN_OUT
      saved_status : "Connection_Status.UDT";
      status_timer : TOF_TIME;
   END_VAR
BEGIN
   "Disconnect_Status.Save_Status"(block_status := #block_status,
                                   saved_status := #saved_status,
                                   status_timer := #status_timer);
   "Disconnect_Status.Clear_Status"(requests := #requests,
                                    saved_status := #saved_status);
END_FUNCTION

FUNCTION "Disconnect_Status.Clear_Status" : Void   // FC163, SCL
{ S7_Optimized_Access := 'TRUE' }
VERSION : 0.1
   VAR_INPUT
      requests : "Connection_Requests.UDT";
   END_VAR
   VAR_IN_OUT
      saved_status : "Connection_Status.UDT";
   END_VAR
BEGIN
   IF #requests.connect THEN
       #saved_status.status := 0;
   END_IF;
END_FUNCTION

// folder: tcpip_connection/requests

FUNCTION_BLOCK "Connection.Request_Disconnect"   // FB1, SCL
{ S7_Optimized_Access := 'TRUE' }
VERSION : 0.1
   VAR_IN_OUT
      hmi : "Connection_Status_Element.UDT";
      sign : "Connection_Requests.UDT";
   END_VAR
   VAR
      _old : Bool;
   END_VAR
BEGIN
   IF "Bool.Falling_Edge"(signal := #hmi.operation_button_actuate, old_signal := #_old) THEN
       #sign.disconnect := TRUE;
   END_IF;
   #_old := #hmi.operation_button_actuate;
END_FUNCTION_BLOCK

FUNCTION_BLOCK "Connection.Requests"   // FB3, SCL
{ S7_Optimized_Access := 'TRUE' }
VERSION : 0.1
   VAR_IN_OUT
      hmi : "Connection_Status_Table.UDT";
      sign : "Connection_Requests.UDT";
   END_VAR
   VAR
      Request_Connect : "Connection.Request_Connect";
      Request_Disconnect : "Connection.Request_Disconnect";
      Request_Send : "Connection.Request_Send";
   END_VAR
BEGIN
   #Request_Connect(hmi := #hmi.connect,
                    sign := #sign);
   #Request_Disconnect(hmi := #hmi.disconnect,
                       sign := #sign);
   #Request_Send(hmi := #hmi.send,
                 sign := #sign);
END_FUNCTION_BLOCK

FUNCTION_BLOCK "Connection.Request_Connect"   // FB4, SCL
{ S7_Optimized_Access := 'TRUE' }
VERSION : 0.1
   VAR_IN_OUT
      hmi : "Connection_Status_Element.UDT";
      sign : "Connection_Requests.UDT";
   END_VAR
   VAR
      _old : Bool;
   END_VAR
BEGIN
   IF "Bool.Falling_Edge"(signal := #hmi.operation_button_actuate, old_signal := #_old) THEN
       #sign.connect := TRUE;
   END_IF;
   #_old := #hmi.operation_button_actuate;
END_FUNCTION_BLOCK

FUNCTION_BLOCK "Connection.Request_Send"   // FB8, SCL
{ S7_Optimized_Access := 'TRUE' }
VERSION : 0.1
   VAR_IN_OUT
      hmi : "Connection_Status_Element.UDT";
      sign : "Connection_Requests.UDT";
   END_VAR
   VAR
      _old : Bool;
   END_VAR
BEGIN
   IF "Bool.Falling_Edge"(signal := #hmi.operation_button_actuate, old_signal := #_old) THEN
       #sign.send := TRUE;
   END_IF;
   #_old := #hmi.operation_button_actuate;
END_FUNCTION_BLOCK

// folder: tcpip_connection/reset

FUNCTION_BLOCK "Reset"   // FB12, SCL
{ S7_Optimized_Access := 'TRUE' }
VERSION : 0.1
   VAR_INPUT
      tcon_param : TCON_Param;
   END_VAR
   VAR_IN_OUT
      requests : "Connection_Requests.UDT";
   END_VAR
   VAR
      T_RESET : T_RESET;
   END_VAR
BEGIN
   #T_RESET(REQ:=#requests.reset,
            ID:=#tcon_param.ID);
   #requests.reset := FALSE;
END_FUNCTION_BLOCK

// folder: tcpip_connection/send

FUNCTION_BLOCK "Send"   // FB9, SCL
{ S7_Optimized_Access := 'TRUE' }